
screen "704_Line_Overview_4" 1280x800
   Button "Button_19" at 852,670 size 37x32; TextOff 'Text'
      on Release: ActivateScreen("711_CARRIER_STATUS", 0)
      on Press: SetTag("HMI_EMS_Nr", "CarrierNumber")
   Button "Template_Button_3" at 1074,2 size 203x55; TextOn 'FAULT RESET FAULT RESET'; TextOff 'FAULT RESET FAULT RESET'
      on Release: ResetBit("DB_SDC_GLOBAL_M.SDC_ER_Reset")
      on Press: SetBit("DB_SDC_GLOBAL_M.SDC_ER_Reset")
   AlarmView "Template_Alarm view_2" at 128,2 size 948x112
   Button "Template_Button_4" at 1196,56 size 81x59; TextOff 'Text'
      Appearance <- "AlwaysTRUE"
   Button "Button_7" at 0,57 size 128x58; TextOff 'SELECT SCREEN'
      on Release: ActivateScreen("010_START", 0)
   Button "Button_6" at 0,0 size 128x58; TextOff 'PREVIOUS SCREEN'
      on Click: function_efd93a16()
   DateTimeField "Template_Date/time field_2" at 1075,56 size 123x28
   DateTimeField "Template_Date/time field_3" at 1075,83 size 122x32
   TextField "Text field_2" at 485,123 size 327x28; Text 'OVERVIEW 4 - SCREEN 704'
   GraphicView "Graphic view_1" at 439,169 size 432x627; Picture "Graphic_4"
   TextField "Text field_34" at 898,673 size 46x25; Text 'S34'
   TextField "Text field_93" at 584,373 size 60x24; Text 'EMS01'
   TextField "Text field_95" at 578,408 size 71x22; Text 'AREA E'
   Button "Button_2" at 988,687 size 127x87; TextOn 'LINE_OVERVIEW_2 LINE OVERVIEW_2'; TextOff 'LINE_OVERVIEW_2 System Overview Screen'
      on Click: ActivateScreen("700_System_Line_Overview", 0)
   Button "Button_1" at 1125,687 size 127x87; TextOn 'LINE_OVERVIEW_2 LINE OVERVIEW_2'; TextOff 'LINE_OVERVIEW_2 / Main Screen'
      on Click: ActivateScreen("010_START", 0)
   Button "Button_3" at 852,182 size 37x32; TextOff 'Text'
      on Release: ActivateScreen("711_CARRIER_STATUS", 0)
      on Press: SetTag("HMI_EMS_Nr", "CarrierNumber")
   Button "Button_4" at 852,215 size 37x32; TextOff 'Text'
      on Release: ActivateScreen("711_CARRIER_STATUS", 0)
      on Press: SetTag("HMI_EMS_Nr", "CarrierNumber")
   Button "Button_5" at 852,250 size 37x32; TextOff 'Text'
      on Release: ActivateScreen("711_CARRIER_STATUS", 0)
      on Press: SetTag("HMI_EMS_Nr", "CarrierNumber")
   Button "Button_8" at 852,285 size 37x32; TextOff 'Text'
      on Release: ActivateScreen("711_CARRIER_STATUS", 0)
      on Press: SetTag("HMI_EMS_Nr", "CarrierNumber")
   Button "Button_9" at 852,320 size 37x32; TextOff 'Text'
      on Release: ActivateScreen("711_CARRIER_STATUS", 0)
      on Press: SetTag("HMI_EMS_Nr", "CarrierNumber")
   Button "Button_10" at 852,355 size 37x32; TextOff 'Text'
      on Release: ActivateScreen("711_CARRIER_STATUS", 0)
      on Press: SetTag("HMI_EMS_Nr", "CarrierNumber")
   Button "Button_11" at 852,390 size 37x32; TextOff 'Text'
      on Release: ActivateScreen("711_CARRIER_STATUS", 0)
      on Press: SetTag("HMI_EMS_Nr", "CarrierNumber")
   Button "Button_12" at 852,425 size 37x32; TextOff 'Text'
      on Release: ActivateScreen("711_CARRIER_STATUS", 0)
      on Press: SetTag("HMI_EMS_Nr", "CarrierNumber")
   Button "Button_13" at 852,460 size 37x32; TextOff 'Text'
      on Release: ActivateScreen("711_CARRIER_STATUS", 0)
      on Press: SetTag("HMI_EMS_Nr", "CarrierNumber")
   Button "Button_14" at 852,495 size 37x32; TextOff 'Text'
      on Release: ActivateScreen("711_CARRIER_STATUS", 0)
      on Press: SetTag("HMI_EMS_Nr", "CarrierNumber")
   Button "Button_15" at 852,530 size 37x32; TextOff 'Text'
      on Release: ActivateScreen("711_CARRIER_STATUS", 0)
      on Press: SetTag("HMI_EMS_Nr", "CarrierNumber")
   Button "Button_16" at 852,565 size 37x32; TextOff 'Text'
      on Release: ActivateScreen("711_CARRIER_STATUS", 0)
      on Press: SetTag("HMI_EMS_Nr", "CarrierNumber")
   Button "Button_17" at 852,600 size 37x32; TextOff 'Text'
      on Release: ActivateScreen("711_CARRIER_STATUS", 0)
      on Press: SetTag("HMI_EMS_Nr", "CarrierNumber")
   Button "Button_18" at 852,635 size 37x32; TextOff 'Text'
      on Release: ActivateScreen("711_CARRIER_STATUS", 0)
      on Press: SetTag("HMI_EMS_Nr", "CarrierNumber")
   IOField "I/O field_50" at 852,670 size 37x32; FormatPattern 99
      ProcessValue <- "CarrierNumber"
      Appearance <- "Faulted"
   IOField "I/O field_32" at 852,182 size 37x32; FormatPattern 99
      ProcessValue <- "CarrierNumber"
      Appearance <- "Faulted"
   IOField "I/O field_33" at 852,215 size 37x32; FormatPattern 99
      ProcessValue <- "CarrierNumber"
      Appearance <- "Faulted"
   IOField "I/O field_34" at 852,250 size 37x32; FormatPattern 99
      ProcessValue <- "CarrierNumber"
      Appearance <- "Faulted"
   IOField "I/O field_35" at 852,285 size 37x32; FormatPattern 99
      ProcessValue <- "CarrierNumber"
      Appearance <- "Faulted"
   IOField "I/O field_36" at 852,320 size 37x32; FormatPattern 99
      ProcessValue <- "CarrierNumber"
      Appearance <- "Faulted"
   IOField "I/O field_49" at 852,635 size 37x32; FormatPattern 99
      ProcessValue <- "CarrierNumber"
      Appearance <- "Faulted"
   IOField "I/O field_40" at 852,600 size 37x32; FormatPattern 99
      ProcessValue <- "CarrierNumber"
      Appearance <- "Faulted"
   IOField "I/O field_41" at 852,565 size 37x32; FormatPattern 99
      ProcessValue <- "CarrierNumber"
      Appearance <- "Faulted"
   IOField "I/O field_43" at 852,530 size 37x32; FormatPattern 99
      ProcessValue <- "CarrierNumber"
      Appearance <- "Faulted"
   IOField "I/O field_44" at 852,495 size 37x32; FormatPattern 99
      ProcessValue <- "CarrierNumber"
      Appearance <- "Faulted"
   IOField "I/O field_45" at 852,460 size 37x32; FormatPattern 99
      ProcessValue <- "CarrierNumber"
      Appearance <- "Faulted"
   IOField "I/O field_46" at 852,425 size 37x32; FormatPattern 99
      ProcessValue <- "CarrierNumber"
      Appearance <- "Faulted"
   IOField "I/O field_47" at 852,390 size 37x32; FormatPattern 99
      ProcessValue <- "CarrierNumber"
      Appearance <- "Faulted"
   IOField "I/O field_48" at 852,355 size 37x32; FormatPattern 99
      ProcessValue <- "CarrierNumber"
      Appearance <- "Faulted"

screen "711_CARRIER_STATUS" 1280x800, template "Top_Header"
   on GenerateScreen: "SDC_EMS_STATUS"("HMI_EMS_Nr"); "SDC_EMS_TA_STATUS"("HMI_EMS_Nr"); "SDC_ERRORS"("HMI_EMS_Nr"); SetTag("SDC\DB_SDC_EMS\HMI[XX].BILD_Nr", 711); SetTag("SDC\_intern_Bildnummer", 711); "SDC_TS_REFERENCE"("SDC\DB_SDC_EMS\EMS[XXX].TS_STAT.VAL.SEK"); "SDC_GLOBAL_REFERENCE_PROFIL"("SDC\DB_SDC_EMS\EMS[XXX].PROFIL")
   on ClearScreen: SetTag("SDC\DB_SDC_EMS\HMI[XX].BILD_Nr", 0)
   IOField "EA-Feld_4" at 270,148 size 56x32; FormatPattern 99
      on OnFinishInput: "SDC_EMS_STATUS"("HMI_EMS_Nr"); "SDC_EMS_TA_STATUS"("HMI_EMS_Nr"); "SDC_ERRORS"("HMI_EMS_Nr")
      ProcessValue <- "HMI_EMS_Nr"
   TextField "Textfeld_3" at 378,151 size 118x25; Text 'EMS-No. / EMS-Number / Carrier-Number'
   Button "Schaltfläche_1" at 327,149 size 40x32; TextOff '+'
      on Click: function_dd21b452("HMI_EMS_Nr", 1); "SDC_EMS_STATUS"("HMI_EMS_Nr"); "SDC_EMS_TA_STATUS"("HMI_EMS_Nr"); "SDC_ERRORS"("HMI_EMS_Nr")
   Button "Schaltfläche_3" at 231,148 size 39x32; TextOff '-'
      on Click: function_b9b71300("HMI_EMS_Nr", 1); "SDC_EMS_STATUS"("HMI_EMS_Nr"); "SDC_EMS_TA_STATUS"("HMI_EMS_Nr"); "SDC_ERRORS"("HMI_EMS_Nr")
   IOField "EA-Feld_5" at 740,309 size 96x32; Authorization "Benutzerverwaltung"; FormatPattern 99999
      ProcessValue <- "HMI_Carrier_ActualSpeed"
   TextField "Textfeld_4" at 706,289 size 187x25; Text 'drive stop position [mm] / Drive Stopposition mm / Current Carrier Speed'
   Group "Gruppe" at 176,202 size 1068x49
   IOField "EA-Feld_14" at 788,216 size 48x28; FormatPattern 999
      on OnFinishInput: "SDC_EMS_STATUS"("HMI_EMS_Nr"); "SDC_TS_REFERENCE"("SDC\DB_SDC_EMS\EMS[XXX].TS_STAT.VAL.SEK"); "SDC_EMS_TA_STATUS"("HMI_EMS_Nr"); "SDC_ERRORS"("HMI_EMS_Nr")
      ProcessValue <- "HMI_EMS_Nr"
   IOField "EA-Feld_15" at 788,216 size 48x28; FormatPattern 999
      on OnFinishInput: "SDC_TS_PARAMETER"()
      Visibility <- "SDC\DB_SDC_EMS\EMS[XXX].TS_STAT.VAL.ERROR"
      ProcessValue <- "DB401_HMI_Status_CarrierFaultCode"
   TextField "Textfeld_17" at 726,216 size 50x22; Text 'ERROR / Error'
      Visibility <- "SDC\DB_SDC_EMS\EMS[XXX].ERRORS_SDC"
   IOField "EA-Feld_22" at 754,168 size 96x32; Authorization "Benutzerverwaltung"; FormatPattern 9999999999
      ProcessValue <- "HMI_Carrier_CurrentPosition"
   TextField "Textfeld_26" at 736,150 size 175x25; Text 'drive in position / Drive in Position / Current carrier position'
   TextField "Textfeld_29" at 1028,255 size 200x25; Text 'distance to next EMS / distance to preceding EMS / Next Stop Position'
   TextField "Textfeld_47" at 452,266 size 177x25; Text 'drives forward / EMS move forward / Carrier Moving Forward'
   Circle "Kreis_22" at 431,272 size 15x15
      Appearance <- "HMI_Carrier_RunningFwd"
   TextField "Textfeld_55" at 452,288 size 176x25; Text 'drives backward / EMS move reward / Carrier Moving Reverse'
   Circle "Kreis_30" at 431,294 size 15x15
      Appearance <- "HMI_Carrier_RunningRev"
   TextField "Textfeld_56" at 452,309 size 179x25; Text 'drive in position / EMS Drive in Position / Carrier Drive in Position'
   Circle "Kreis_31" at 431,315 size 15x15
      Appearance <- "HMI_Carrier_AtCommandPosition"
   Button "Schaltfläche_15" at 11,710 size 117x84; TextOff 'I / O EDIT CARRIER I/O'
      on Click: ActivateScreen("712_CARRIER_IO", 0)
   TextField "Textfeld_7" at 567,118 size 243x27; Text 'section counter / min Barcode mm / Carrier Status'
   Rectangle "Rectangle_1" at 11,443 size 55x42
      Appearance <- "HMI_Carrier_DriveCommFault"
   TextField "Textfeld_8" at 71,450 size 155x25; Text 'EMS Notbetrieb Tilt / EMS VAC CLEAN / G120 D Drive Status'
   Rectangle "Rectangle_2" at 11,494 size 55x42
      Appearance <- "HMI_Carrier_EncoderCommFault"
   TextField "Textfeld_9" at 74,501 size 148x25; Text 'EMS Notbetrieb Tilt / EMS VAC CLEAN / PnF Encoder Status'
   Rectangle "Rectangle_9" at 11,547 size 55x42
      Appearance <- "HMI_Carrier_HMICommFault"
   TextField "Textfeld_16" at 76,552 size 152x25; Text 'EMS Notbetrieb Tilt / EMS VAC CLEAN / IRD 400 HMI Status'
   TextField "Textfeld_19" at 12,400 size 242x26; Text 'EMS Notbetrieb Tilt / EMS VAC CLEAN / CARRIER DEVICE STATUS'
   Button "Schaltfläche_2" at 546,476 size 27x27; TextOff 'Text'; Authorization "Bedienen"
      on Click: function_c82f6f27("SDC\DB_SDC_EMS\EMS[XXX].FKT_SET", 8)
      ObjectEnable <- "SDC\DB_SDC_EMS\HMI[XX].FR_EDIT"
      Appearance <- "HMI_Carrier_Comm_Fault"
   Button "Schaltfläche_5" at 546,506 size 27x27; TextOff 'Text'; Authorization "Bedienen"
      on Click: function_c82f6f27("SDC\DB_SDC_EMS\EMS[XXX].FKT_SET", 10)
      ObjectEnable <- "SDC\DB_SDC_EMS\HMI[XX].FR_EDIT"
      Appearance <- "HMI_Carrier_Auto"
   Button "Schaltfläche_6" at 546,566 size 27x27; TextOff 'Text'; Authorization "Bedienen"
      on Click: function_c82f6f27("SDC\DB_SDC_EMS\EMS[XXX].FKT_SET", 12)
      ObjectEnable <- "SDC\DB_SDC_EMS\HMI[XX].FR_EDIT"
      Appearance <- "HMI_Carrier_Faulted"
   Button "Schaltfläche_7" at 546,596 size 27x27; TextOff 'Text'; Authorization "Bedienen"
      on Click: function_c82f6f27("SDC\DB_SDC_EMS\EMS[XXX].FKT_SET", 13)
      ObjectEnable <- "SDC\DB_SDC_EMS\HMI[XX].FR_EDIT"
      Appearance <- "HMI_Carrier_HoldPBPressed"
   Button "Schaltfläche_9" at 546,536 size 27x27; TextOff 'Text'; Authorization "Bedienen"
      on Click: function_c82f6f27("SDC\DB_SDC_EMS\EMS[XXX].FKT_SET", 11)
      ObjectEnable <- "SDC\DB_SDC_EMS\HMI[XX].FR_EDIT"
      Appearance <- "HMI_Carrier_Manual"
   TextField "Textfeld_59" at 579,598 size 176x25; Text 'Kohle Test n.i.O. / EMS TO REPAIR / CARRIER PROD. HOLD'
   TextField "Textfeld_1" at 579,507 size 148x25; Text 'EMS Notbetrieb Tilt / EMS VAC CLEAN / CARRIER IN AUTO'
   TextField "Textfeld_2" at 579,568 size 159x25; Text 'SMGM Qualität n.i.O. / EMS TO REPAIR / CARRIER FAULT'
   TextField "Textfeld_20" at 580,476 size 181x25; Text 'EMS Notbetrieb Tilt / EMS VAC CLEAN / CARRIER COMM FAULT'
   TextField "Textfeld_6" at 580,536 size 166x25; Text 'EMS Notbetrieb Tilt / EMS VAC CLEAN / CARRIER IN MANUAL'
   TextField "Textfeld_38" at 218,274 size 188x25; Text 'command drive forward / Command forward / Command Drive Forward'
   Circle "Kreis_13" at 194,280 size 15x15
      Appearance <- "HMI_Carrier_DriveFwdCommand"
   TextField "Textfeld_40" at 218,305 size 193x25; Text 'command drive backward / Command reward / Command Speed'
   IOField "EA-Feld_1" at 138,302 size 96x32; Authorization "Benutzerverwaltung"; FormatPattern 99999
      ProcessValue <- "HMI_Carrier_DriveCmdSpeed"
   Button "Schaltfläche_10" at 154,710 size 117x84; TextOff 'I / O EDIT CARRIER DRIVE'
      on Click: ActivateScreen("728_CARRIER_VFD_STATUS", 0)
   Button "Schaltfläche_11" at 300,710 size 117x84; TextOff 'I / O EDIT CARRIER FAULTS'
      on Click: ActivateScreen("713_CARRIER_FAULT", 0)
   IOField "EA-Feld_2" at 1116,273 size 96x32; Authorization "Benutzerverwaltung"; FormatPattern 99999999
      ProcessValue <- "HMI_Carrier_NextStopPosition"
   TextField "Textfeld_11" at 1030,147 size 200x25; Text 'distance to next EMS / distance to preceding EMS / Next Carrier Number'
   IOField "EA-Feld_3" at 1118,165 size 96x32; Authorization "Benutzerverwaltung"; FormatPattern 99999
      ProcessValue <- "HMI_Carrier_NextCarrierNumber"
   IOField "EA-Feld_30" at 951,487 size 56x32; FormatPattern 99
      on OnFinishInput: "SDC_TS_PARAMETER"()
      ProcessValue <- "HMI_Carrier_CurrentZone"
   TextField "Textfeld_37" at 825,487 size 174x27; Text 'section no. / Tracksectionnumber / Zone Number'
   TextField "Textfeld_5" at 825,466 size 174x27; Text 'section no. / Tracksectionnumber / Carrier in'
   Button "Schaltfläche_4" at 1089,543 size 117x84; TextOff 'I / O EDIT SET MASK CARRIER FAULTS'
      Appearance <- "Mask_Carrier_Faults_LT"
      on Press: SetBit("Set_Mask_Carrier_Faults_PB")
      on Release: ResetBit("Set_Mask_Carrier_Faults_PB")
   Button "Schaltfläche_8" at 1089,670 size 117x84; TextOff 'I / O EDIT RESET MASK CARRIER FAULTS'
      on Press: SetBit("Reset_Mask_Carrier_Faults_PB")
      on Release: ResetBit("Reset_Mask_Carrier_Faults_PB")
   IOField "EA-Feld_6" at 951,552 size 56x32; FormatPattern ??
      on OnFinishInput: "SDC_TS_PARAMETER"()
      ProcessValue <- "HMI_Carrier_CurrentArea"
   TextField "Textfeld_10" at 825,552 size 174x27; Text 'section no. / Tracksectionnumber / Area Number'
   TextField "Textfeld_12" at 825,531 size 174x27; Text 'section no. / Tracksectionnumber / Carrier in'

screen "713_CARRIER_FAULT" 1280x800, template "Top_Header"
   on GenerateScreen: "SDC_EMS_STATUS"('SDC\_EMS_Nr'); "SDC_TS_REFERENCE"("SDC\_TS_Nr"); SetTag("SDC\_intern_Bildnummer", 712); "SDC_EMS_TA_STATUS"("HMI_EMS_Nr"); SetTag("SDC\_intern_Bildnummer", 712)
   on ClearScreen: SetTag("SDC\DB_SDC_EMS\HMI[XX].BILD_Nr", 0)
   IOField "EA-Feld_4" at 510,185 size 56x32; FormatPattern 9999
      on OnFinishInput: "SDC_EMS_STATUS"("HMI_EMS_Nr"); "SDC_EMS_TA_STATUS"("HMI_EMS_Nr"); "SDC_ERRORS"("HMI_EMS_Nr")
      ProcessValue <- "HMI_EMS_Nr"
   TextField "Textfeld_3" at 618,188 size 118x25; Text 'EMS-No. / EMS-Number / Carrier-Number'
   Button "Schaltfläche_1" at 567,185 size 40x32; TextOff '+'
      on Click: function_dd21b452("HMI_EMS_Nr", 1); "SDC_EMS_STATUS"("HMI_EMS_Nr"); "SDC_EMS_TA_STATUS"("HMI_EMS_Nr"); "SDC_ERRORS"("HMI_EMS_Nr")
   Button "Schaltfläche_3" at 470,185 size 39x32; TextOff '-'
      on Click: function_b9b71300("HMI_EMS_Nr", 1); "SDC_EMS_STATUS"("HMI_EMS_Nr"); "SDC_EMS_TA_STATUS"("HMI_EMS_Nr"); "SDC_ERRORS"("HMI_EMS_Nr")
   TextField "Textfeld_7" at 550,118 size 243x27; Text 'section counter / min Barcode mm / Carrier Fault'
   Button "Button_1" at 84,303 size 50x246; TextOff 'Text'
   TextField "Textfeld_11" at 137,309 size 293x25; Text 'EMS-No. / EMS-Number / FAULT 01 - CARRIER GENERAL FAULT'
   TextField "Textfeld_10" at 137,335 size 238x25; Text 'EMS-No. / EMS-Number / FAULT 02 - MOTION ON FAULT'
   TextField "Textfeld_13" at 137,361 size 245x25; Text 'EMS-No. / EMS-Number / FAULT 03 - MOTION OFF FAULT'
   TextField "Textfeld_14" at 137,387 size 288x25; Text 'EMS-No. / EMS-Number / FAULT 04 - CARRIER SPACING FAULT'
   TextField "Textfeld_15" at 137,412 size 248x25; Text 'EMS-No. / EMS-Number / FAULT 05 - DRIVE COMM FAULT'
   TextField "Textfeld_16" at 137,438 size 272x25; Text 'EMS-No. / EMS-Number / FAULT 06 - DRIVE GENERAL FAULT'
   TextField "Textfeld_17" at 137,464 size 275x25; Text 'EMS-No. / EMS-Number / FAULT 07 - ENCODER COMM FAULT'
   TextField "Textfeld_18" at 137,490 size 265x25; Text 'EMS-No. / EMS-Number / FAULT 08 - CRASH DETECT FAULT'
   Circle "Kreis_13" at 102,312 size 15x15
      Appearance <- "DB401_HMI_Status_CarrierFaultCode"
   Circle "Kreis_1" at 102,338 size 15x15
      Appearance <- "DB401_HMI_Status_CarrierFaultCode"
   Circle "Kreis_2" at 102,364 size 15x15
      Appearance <- "DB401_HMI_Status_CarrierFaultCode"
   Circle "Kreis_3" at 102,390 size 15x15
      Appearance <- "DB401_HMI_Status_CarrierFaultCode"
   Circle "Kreis_4" at 102,416 size 15x15
      Appearance <- "DB401_HMI_Status_CarrierFaultCode"
   Circle "Kreis_5" at 102,442 size 15x15
      Appearance <- "DB401_HMI_Status_CarrierFaultCode"
   Circle "Kreis_6" at 102,468 size 15x15
      Appearance <- "DB401_HMI_Status_CarrierFaultCode"
   Circle "Kreis_7" at 102,494 size 15x15
      Appearance <- "DB401_HMI_Status_CarrierFaultCode"
   TextField "Textfeld_1" at 137,516 size 337x25; Text 'EMS-No. / EMS-Number / FAULT 15 - DRIVE ERROR INTERNAL COMM'
   Circle "Kreis_8" at 102,520 size 15x15
      Appearance <- "DB401_HMI_Status_CarrierFaultCode"
   Button "Button_2" at 516,303 size 50x246; TextOff 'Text'
   TextField "Textfeld_2" at 569,309 size 326x25; Text 'EMS-No. / EMS-Number / FAULT 20 - DRIVE MOTOR OVERCURRENT'
   TextField "Textfeld_4" at 569,335 size 273x25; Text 'EMS-No. / EMS-Number / FAULT 23 - DRIVE UNDERVOLTAGE'
   TextField "Textfeld_5" at 569,361 size 261x25; Text 'EMS-No. / EMS-Number / FAULT 24 - DRIVE OVERVOLTAGE'
   TextField "Textfeld_6" at 569,387 size 349x25; Text 'EMS-No. / EMS-Number / FAULT 25 - DRIVE PWR MODULE NOT READY'
   TextField "Textfeld_8" at 569,412 size 294x25; Text 'EMS-No. / EMS-Number / FAULT 32 - DRIVE MOTOR OVERTEMP'
   TextField "Textfeld_9" at 569,438 size 302x25; Text 'EMS-No. / EMS-Number / FAULT 40 - CARRIER NUMBER INVALID'
   TextField "Textfeld_12" at 569,464 size 302x25; Text 'EMS-No. / EMS-Number / FAULT 60 - ENCODER POSITION FAULT'
   Circle "Kreis_9" at 534,312 size 15x15
      Appearance <- "DB401_HMI_Status_CarrierFaultCode"
   Circle "Kreis_10" at 534,338 size 15x15
      Appearance <- "DB401_HMI_Status_CarrierFaultCode"
   Circle "Kreis_11" at 534,364 size 15x15
      Appearance <- "DB401_HMI_Status_CarrierFaultCode"
   Circle "Kreis_12" at 534,390 size 15x15
      Appearance <- "DB401_HMI_Status_CarrierFaultCode"
   Circle "Kreis_14" at 534,416 size 15x15
      Appearance <- "DB401_HMI_Status_CarrierFaultCode"
   Circle "Kreis_15" at 534,442 size 15x15
      Appearance <- "DB401_HMI_Status_CarrierFaultCode"
   Circle "Kreis_16" at 534,468 size 15x15
      Appearance <- "DB401_HMI_Status_CarrierFaultCode"
   TextField "Textfeld_20" at 569,489 size 339x25; Text 'EMS-No. / EMS-Number / FAULT DUP - DUPLICATE CARRIER # FAULT'
   Circle "Kreis_18" at 534,493 size 15x15
      Appearance <- "DB401_HMI_Status_CarrierFaultCode"

screen "715_ACCESS_POINT_LAYOUT" 1280x800
   GraphicView "Graphic view_1" at 0,119 size 1144x681; Picture "LAYOUT 1"
   Button "Button_9" at 451,171 size 47x26; TextOff 'AP6'
      Appearance <- "[106]"
   Button "Button_12" at 517,123 size 46x26; TextOff 'AP7'
      Appearance <- "[107]"
   Button "Button_10" at 574,123 size 46x26; TextOff 'AP8'
      Appearance <- "[108]"
   Button "Button_11" at 627,123 size 45x26; TextOff 'AP9'
      Appearance <- "[109]"
   Button "Button_13" at 694,171 size 47x26; TextOff 'AP5'
      Appearance <- "[105]"
   Button "Button_8" at 734,123 size 50x26; TextOff 'AP10'
      Appearance <- "[110]"
   Button "Button_14" at 749,222 size 52x26; TextOff 'AP11'
      Appearance <- "[111]"
   Button "Button_7" at 750,325 size 51x26; TextOff 'AP4'
      Appearance <- "[104]"
   Button "Button_6" at 749,444 size 52x26; TextOff 'AP12'
      Appearance <- "[112]"
   Button "Button_5" at 751,607 size 51x26; TextOff 'AP3'
      Appearance <- "[103]"
   Button "Button_4" at 777,637 size 52x26; TextOff 'AP13'
      Appearance <- "[113]"
   Button "Button_15" at 576,726 size 52x26; TextOff 'AP14'
      Appearance <- "[114]"
   Button "Button_16" at 384,711 size 53x26; TextOff 'AP15'
      Appearance <- "[115]"
   Button "Button_17" at 295,743 size 52x26; TextOff 'AP16'
      Appearance <- "[116]"
   Button "Button_18" at 267,687 size 53x26; TextOff 'AP17'
      Appearance <- "[117]"
   Button "Button_19" at 329,611 size 51x26; TextOff 'AP18'
      Appearance <- "[118]"
   Button "Button_1" at 479,611 size 50x26; TextOff 'AP1'
      Appearance <- "[101]"
   Button "Button_2" at 620,612 size 50x26; TextOff 'AP2'
      Appearance <- "[102]"
   TextField "Text field_126" at 847,138 size 369x28; Text 'ACCESS POINT LAYOUT SCREEN'
   Button "Button_20" at 471,117 size 46x26; TextOff 'AP19'
      Appearance <- "[119]"
   Button "Template_Button_3" at 1074,2 size 203x55; TextOn 'FAULT RESET FAULT RESET'; TextOff 'FAULT RESET FAULT RESET'
      on Release: ResetBit("DB_SDC_GLOBAL_M.SDC_ER_Reset")
      on Press: SetBit("DB_SDC_GLOBAL_M.SDC_ER_Reset")
   AlarmView "Template_Alarm view_2" at 128,2 size 948x112
   Button "Template_Button_4" at 1196,56 size 81x59; TextOff 'Text'
      Appearance <- "AlwaysTRUE"
   Button "Button_21" at 0,57 size 128x58; TextOff 'SELECT SCREEN'
      on Release: ActivateScreen("010_START", 0)
   Button "Button_22" at 0,0 size 128x58; TextOff 'PREVIOUS SCREEN'
      on Click: function_efd93a16()
   DateTimeField "Template_Date/time field_2" at 1075,56 size 123x28
   DateTimeField "Template_Date/time field_3" at 1075,83 size 122x32

screen "708_ZONE_STATUS" 1280x800, template "Top_Header"
   on GenerateScreen: "SDC_TS_PARAMETER"(); "SDC_TS_REFERENCE"("HMI_Zone_Nr"); SetTag("SDC\DB_SDC_TS_PARAMETER\DB_SDC_TS_PARAMETER_HMI.HMI[XX].BILD_Nr", 704); SetTag("SDC\_intern_Bildnummer", 704)
   on ClearScreen: SetTag("SDC\DB_SDC_TS_PARAMETER\DB_SDC_TS_PARAMETER_HMI.HMI[XX].BILD_Nr", 0)
   IOField "EA-Feld_1" at 144,392 size 96x32; Authorization "Benutzerverwaltung"; FormatPattern 9999999999
      Appearance <- "SDC\DB_SDC_TS_PARAMETER\DB_SDC_TS_PARAMETER_HMI.HMI[XX].FR_EDIT"
      ObjectEnable <- "SDC\DB_SDC_TS_PARAMETER\DB_SDC_TS_PARAMETER_HMI.HMI[XX].FR_EDIT"
      ProcessValue <- "DB401_HMI_Status_ZoneStatus.ZoneStartPosition"
   TextField "Textfeld_1" at 137,344 size 272x58; Text 'barcode value at start of section [mm] Sektion Start Barcode mm Position at start of zone [mm]'
   IOField "EA-Feld_2" at 1022,324 size 96x32; Authorization "Benutzerverwaltung"; FormatPattern 9999999999
      Appearance <- "SDC\DB_SDC_TS_PARAMETER\DB_SDC_TS_PARAMETER_HMI.HMI[XX].FR_EDIT"
      ObjectEnable <- "SDC\DB_SDC_TS_PARAMETER\DB_SDC_TS_PARAMETER_HMI.HMI[XX].FR_EDIT"
      ProcessValue <- "DB401_HMI_Status_ZoneStatus.ZoneEndPosition"
   TextField "Textfeld_2" at 743,318 size 275x59; Text 'barcode value at end of section [mm] Sektion Ende Barcode mm Position at end of zone [mm]'
   IOField "EA-Feld_4" at 416,188 size 56x32; FormatPattern 9999
      on OnFinishInput: "SDC_TS_PARAMETER"(); "SDC_TS_REFERENCE"("HMI_Zone_Nr")
      ProcessValue <- "HMI_Zone_Nr"
   TextField "Textfeld_3" at 515,188 size 93x33; Text 'section no. / Sektionnumber / Zone No'
   Button "Schaltfläche_1" at 473,188 size 40x32; TextOff '+'
      on Click: function_dd21b452("HMI_Zone_Nr", 1); "SDC_TS_PARAMETER"(); "SDC_TS_REFERENCE"("HMI_Zone_Nr")
   Button "Schaltfläche_3" at 376,188 size 39x32; TextOff '-'
      on Click: function_b9b71300("HMI_Zone_Nr", 1); "SDC_TS_PARAMETER"(); "SDC_TS_REFERENCE"("HMI_Zone_Nr")
   IOField "EA-Feld_8" at 1056,188 size 56x32; Authorization "Benutzerverwaltung"; FormatPattern 9999
      Appearance <- "SDC\DB_SDC_TS_PARAMETER\DB_SDC_TS_PARAMETER_HMI.HMI[XX].FR_EDIT"
      ObjectEnable <- "SDC\DB_SDC_TS_PARAMETER\DB_SDC_TS_PARAMETER_HMI.HMI[XX].FR_EDIT"
      ProcessValue <- "DB401_HMI_Status_ZoneStatus.NextZoneNumber"
   TextField "Textfeld_7" at 957,187 size 107x33; Text 'next section 1 / next Sektion 1 / Next Zone'
   Group "Gruppe" at 141,244 size 1024x49
   IOField "EA-Feld_13" at 610,192 size 163x24; Authorization "Benutzerverwaltung"; FormatPattern ????????????????
      Appearance <- "SDC\DB_SDC_TS_PARAMETER\DB_SDC_TS_PARAMETER_HMI.HMI[XX].FR_EDIT"
      ObjectEnable <- "SDC\DB_SDC_TS_PARAMETER\DB_SDC_TS_PARAMETER_HMI.HMI[XX].FR_EDIT"
      ProcessValue <- "DB401_HMI_Status_ZoneStatus.ZoneType"
   TextField "Textfeld_5" at 658,381 size 330x33; Text 'stop position (offset start) mm / Stopposition (Offset Start) mm / Zone Full'
   TextField "Textfeld_6" at 659,422 size 330x33; Text 'stop position (offset start) mm / Stopposition (Offset Start) mm / Speed Zone'
   TextField "Textfeld_8" at 659,463 size 330x33; Text 'stop position (offset start) mm / Stopposition (Offset Start) mm / Speed Zone Start'
   TextField "Textfeld_9" at 659,504 size 330x33; Text 'stop position (offset start) mm / Stopposition (Offset Start) mm / Speed Zone End'
   IOField "EA-Feld_3" at 596,460 size 56x32; FormatPattern 9999999999
      on OnFinishInput: "SDC_TS_PARAMETER"(); "SDC_TS_REFERENCE"("SDC\_TS_Nr")
      ProcessValue <- "DB401_HMI_Status_ZoneStatus.SpeedZoneStartPos"
   IOField "EA-Feld_6" at 596,500 size 56x32; FormatPattern 9999999999
      on OnFinishInput: "SDC_TS_PARAMETER"(); "SDC_TS_REFERENCE"("SDC\_TS_Nr")
      ProcessValue <- "DB401_HMI_Status_ZoneStatus.SpeedZoneEndPos"
   Circle "Kreis_13" at 616,387 size 15x15
      Appearance <- "DB401_HMI_Status_ZoneStatus.ZoneFull"
   Circle "Kreis_1" at 616,427 size 15x15
      Appearance <- "DB401_HMI_Status_ZoneStatus.SpeedZone"
   IOField "EA-Feld_9" at 596,540 size 56x32; Authorization "Benutzerverwaltung"; FormatPattern 99999
      Appearance <- "SDC\DB_SDC_TS_PARAMETER\DB_SDC_TS_PARAMETER_HMI.HMI[XX].FR_EDIT"
      ObjectEnable <- "SDC\DB_SDC_TS_PARAMETER\DB_SDC_TS_PARAMETER_HMI.HMI[XX].FR_EDIT"
      ProcessValue <- "DB401_HMI_Status_ZoneStatus.AccumZoneSpacing"
   TextField "Textfeld_11" at 659,542 size 330x33; Text 'stop position (offset start) mm / Stopposition (Offset Start) mm / Accum Zone Spacing'
   IOField "EA-Feld_10" at 596,580 size 56x32; Authorization "Benutzerverwaltung"; FormatPattern 99999
      Appearance <- "SDC\DB_SDC_TS_PARAMETER\DB_SDC_TS_PARAMETER_HMI.HMI[XX].FR_EDIT"
      ObjectEnable <- "SDC\DB_SDC_TS_PARAMETER\DB_SDC_TS_PARAMETER_HMI.HMI[XX].FR_EDIT"
      ProcessValue <- "DB401_HMI_Status_ZoneStatus.ProductionZoneSpacing"
   TextField "Textfeld_12" at 659,582 size 330x33; Text 'stop position (offset start) mm / Stopposition (Offset Start) mm / Prooduction Zone Spacing'
   TextField "Textfeld_13" at 459,114 size 243x27; Text 'section counter / min Barcode mm / Zone Status'
   TextField "Text field_1" at 911,358 size 101x25; Text 'Stop Position'
   TextField "Text field_2" at 642,168 size 83x25; Text 'Zone Type'
   IOField "EA-Feld_5" at 119,189 size 56x32; Authorization "Benutzerverwaltung"; FormatPattern 9999
      Appearance <- "SDC\DB_SDC_TS_PARAMETER\DB_SDC_TS_PARAMETER_HMI.HMI[XX].FR_EDIT"
      ObjectEnable <- "SDC\DB_SDC_TS_PARAMETER\DB_SDC_TS_PARAMETER_HMI.HMI[XX].FR_EDIT"
      ProcessValue <- "DB401_HMI_Status_ZoneStatus.PrevZoneNumber"
   TextField "Textfeld_4" at 25,189 size 94x33; Text 'next section 1 / next Sektion 1 / Prev Zone'

VB script "SDC_EMS_FLAGS"
   'HINWEIS:
   ' Beim Erstellen von Skripten können Sie mit <Strg+Leertaste> vordefinierte 
   ' Systemfunktionen in das neue Skript einbinden.
   ' Das HMIRuntime-Objekt ermöglicht einfachen Zugriff auf die Objekte des
   ' WinCC flexible Objektmodells, ihre Methoden und ihre Eigenschaften.
   ' Für ein komfortables Auswählen einer Objektreferenz betätigen Sie bitte <Alt+Rechts>.
   ' Komplexe Skripte können Sie mit Sprachelementen der Programmiersprache
   ' VBScript erstellen.
   ' Der Zugriff auf WinCC flexible Variablen erfolgt direkt über den Variablennamen,
   ' z.B. Tag = 5
   
   '________________________________________________________________________________
   '
   
   ' Groiß Andreas
   ' Siemens AG Österreich 
   ' Linz Kraußstraße 1-7 
   ' RC-AT I-IA AS-FA-SO-AE2
   ' 28.01.2015
   
   Dim EMS_Nr ' Sektion Number
   Dim Laenge_Data ' Länge FLAG Daten
   Dim Allg_Offset ' Allg Parameter Offset
   Dim HMIFlagDaten_Offset ' HMI Sektionsdaten Offset
   Dim HMI_Nr ' HMI Nummer
   
   ' INIT-------------------------------------------------------------
   
   If (SmartTags("SDC\DB_SDC_EMS_FLAGS\_EMS_Nr") < SmartTags("DB_SDC_GLOBAL_EMS_ID_MIN")) Or (SmartTags("SDC\DB_SDC_EMS_FLAGS\_EMS_Nr") > SmartTags("DB_SDC_GLOBAL_EMS_ID_MAX")) Then
   	SmartTags("SDC\DB_SDC_EMS_FLAGS\_EMS_Nr") = 	SmartTags("DB_SDC_GLOBAL_EMS_ID_MIN")
   End If	
   
   If (SmartTags("SDC\DB_SDC_EMS_FLAGS\_EMS_Nr") < 1) Then
   	SmartTags("SDC\DB_SDC_EMS_FLAGS\_EMS_Nr") = 1
   End If	
   
   '##############################################
   ' S7 sucht sich Daten:
   '##############################################
   
       Laenge_Data = SmartTags("DB_SDC_EMS_FLAGS_HEADER.LAENGE_EMS_FLAGS")
       Allg_Offset = SmartTags("DB_SDC_EMS_FLAGS_HEADER.START_EMS")
   
       SmartTags("SDC\DB_SDC_EMS_FLAGS\_EMS_Flags_Byte_EMS001") = 001 * Laenge_Data - Laenge_Data + Allg_Offset 
       SmartTags("SDC\DB_SDC_EMS_FLAGS\_EMS_Flags_Byte_EMS002") = 002 * Laenge_Data - Laenge_Data + Allg_Offset 
       SmartTags("SDC\DB_SDC_EMS_FLAGS\_EMS_Flags_Byte_EMS003") = 003 * Laenge_Data - Laenge_Data + Allg_Offset 
       SmartTags("SDC\DB_SDC_EMS_FLAGS\_EMS_Flags_Byte_EMS004") = 004 * Laenge_Data - Laenge_Data + Allg_Offset 
       SmartTags("SDC\DB_SDC_EMS_FLAGS\_EMS_Flags_Byte_EMS005") = 005 * Laenge_Data - Laenge_Data + Allg_Offset 
       SmartTags("SDC\DB_SDC_EMS_FLAGS\_EMS_Flags_Byte_EMS006") = 006 * Laenge_Data - Laenge_Data + Allg_Offset 
       SmartTags("SDC\DB_SDC_EMS_FLAGS\_EMS_Flags_Byte_EMS007") = 007 * Laenge_Data - Laenge_Data + Allg_Offset 
       SmartTags("SDC\DB_SDC_EMS_FLAGS\_EMS_Flags_Byte_EMS008") = 008 * Laenge_Data - Laenge_Data + Allg_Offset 
       SmartTags("SDC\DB_SDC_EMS_FLAGS\_EMS_Flags_Byte_EMS009") = 009 * Laenge_Data - Laenge_Data + Allg_Offset 
       SmartTags("SDC\DB_SDC_EMS_FLAGS\_EMS_Flags_Byte_EMS010") = 010 * Laenge_Data - Laenge_Data + Allg_Offset 
       SmartTags("SDC\DB_SDC_EMS_FLAGS\_EMS_Flags_Byte_EMS011") = 011 * Laenge_Data - Laenge_Data + Allg_Offset 
       SmartTags("SDC\DB_SDC_EMS_FLAGS\_EMS_Flags_Byte_EMS012") = 012 * Laenge_Data - Laenge_Data + Allg_Offset 
       SmartTags("SDC\DB_SDC_EMS_FLAGS\_EMS_Flags_Byte_EMS013") = 013 * Laenge_Data - Laenge_Data + Allg_Offset 
       SmartTags("SDC\DB_SDC_EMS_FLAGS\_EMS_Flags_Byte_EMS014") = 014 * Laenge_Data - Laenge_Data + Allg_Offset 
       SmartTags("SDC\DB_SDC_EMS_FLAGS\_EMS_Flags_Byte_EMS015") = 015 * Laenge_Data - Laenge_Data + Allg_Offset 
       SmartTags("SDC\DB_SDC_EMS_FLAGS\_EMS_Flags_Byte_EMS016") = 016 * Laenge_Data - Laenge_Data + Allg_Offset 
       SmartTags("SDC\DB_SDC_EMS_FLAGS\_EMS_Flags_Byte_EMS017") = 017 * Laenge_Data - Laenge_Data + Allg_Offset 
       SmartTags("SDC\DB_SDC_EMS_FLAGS\_EMS_Flags_Byte_EMS018") = 018 * Laenge_Data - Laenge_Data + Allg_Offset 
       SmartTags("SDC\DB_SDC_EMS_FLAGS\_EMS_Flags_Byte_EMS019") = 019 * Laenge_Data - Laenge_Data + Allg_Offset 
       SmartTags("SDC\DB_SDC_EMS_FLAGS\_EMS_Flags_Byte_EMS020") = 020 * Laenge_Data - Laenge_Data + Allg_Offset 
       SmartTags("SDC\DB_SDC_EMS_FLAGS\_EMS_Flags_Byte_EMS021") = 021 * Laenge_Data - Laenge_Data + Allg_Offset 
       SmartTags("SDC\DB_SDC_EMS_FLAGS\_EMS_Flags_Byte_EMS022") = 022 * Laenge_Data - Laenge_Data + Allg_Offset 
       SmartTags("SDC\DB_SDC_EMS_FLAGS\_EMS_Flags_Byte_EMS023") = 023 * Laenge_Data - Laenge_Data + Allg_Offset 
       SmartTags("SDC\DB_SDC_EMS_FLAGS\_EMS_Flags_Byte_EMS024") = 024 * Laenge_Data - Laenge_Data + Allg_Offset 
       SmartTags("SDC\DB_SDC_EMS_FLAGS\_EMS_Flags_Byte_EMS025") = 025 * Laenge_Data - Laenge_Data + Allg_Offset 
       SmartTags("SDC\DB_SDC_EMS_FLAGS\_EMS_Flags_Byte_EMS026") = 026 * Laenge_Data - Laenge_Data + Allg_Offset 
       SmartTags("SDC\DB_SDC_EMS_FLAGS\_EMS_Flags_Byte_EMS027") = 027 * Laenge_Data - Laenge_Data + Allg_Offset 
       SmartTags("SDC\DB_SDC_EMS_FLAGS\_EMS_Flags_Byte_EMS028") = 028 * Laenge_Data - Laenge_Data + Allg_Offset 
       SmartTags("SDC\DB_SDC_EMS_FLAGS\_EMS_Flags_Byte_EMS029") = 029 * Laenge_Data - Laenge_Data + Allg_Offset 
       SmartTags("SDC\DB_SDC_EMS_FLAGS\_EMS_Flags_Byte_EMS030") = 030 * Laenge_Data - Laenge_Data + Allg_Offset 
       SmartTags("SDC\DB_SDC_EMS_FLAGS\_EMS_Flags_Byte_EMS031") = 031 * Laenge_Data - Laenge_Data + Allg_Offset 
       SmartTags("SDC\DB_SDC_EMS_FLAGS\_EMS_Flags_Byte_EMS032") = 032 * Laenge_Data - Laenge_Data + Allg_Offset 
       SmartTags("SDC\DB_SDC_EMS_FLAGS\_EMS_Flags_Byte_EMS033") = 033 * Laenge_Data - Laenge_Data + Allg_Offset 
       SmartTags("SDC\DB_SDC_EMS_FLAGS\_EMS_Flags_Byte_EMS034") = 034 * Laenge_Data - Laenge_Data + Allg_Offset 
       SmartTags("SDC\DB_SDC_EMS_FLAGS\_EMS_Flags_Byte_EMS035") = 035 * Laenge_Data - Laenge_Data + Allg_Offset 
       SmartTags("SDC\DB_SDC_EMS_FLAGS\_EMS_Flags_Byte_EMS036") = 036 * Laenge_Data - Laenge_Data + Allg_Offset 
       SmartTags("SDC\DB_SDC_EMS_FLAGS\_EMS_Flags_Byte_EMS037") = 037 * Laenge_Data - Laenge_Data + Allg_Offset 
       SmartTags("SDC\DB_SDC_EMS_FLAGS\_EMS_Flags_Byte_EMS038") = 038 * Laenge_Data - Laenge_Data + Allg_Offset 
       SmartTags("SDC\DB_SDC_EMS_FLAGS\_EMS_Flags_Byte_EMS039") = 039 * Laenge_Data - Laenge_Data + Allg_Offset     
       SmartTags("SDC\DB_SDC_EMS_FLAGS\_EMS_Flags_Byte_EMS040") = 040 * Laenge_Data - Laenge_Data + Allg_Offset 
       SmartTags("SDC\DB_SDC_EMS_FLAGS\_EMS_Flags_Byte_EMS041") = 041 * Laenge_Data - Laenge_Data + Allg_Offset 
       SmartTags("SDC\DB_SDC_EMS_FLAGS\_EMS_Flags_Byte_EMS042") = 042 * Laenge_Data - Laenge_Data + Allg_Offset 
       SmartTags("SDC\DB_SDC_EMS_FLAGS\_EMS_Flags_Byte_EMS043") = 043 * Laenge_Data - Laenge_Data + Allg_Offset 
       SmartTags("SDC\DB_SDC_EMS_FLAGS\_EMS_Flags_Byte_EMS044") = 044 * Laenge_Data - Laenge_Data + Allg_Offset 
       SmartTags("SDC\DB_SDC_EMS_FLAGS\_EMS_Flags_Byte_EMS045") = 045 * Laenge_Data - Laenge_Data + Allg_Offset 
       SmartTags("SDC\DB_SDC_EMS_FLAGS\_EMS_Flags_Byte_EMS046") = 046 * Laenge_Data - Laenge_Data + Allg_Offset 
       SmartTags("SDC\DB_SDC_EMS_FLAGS\_EMS_Flags_Byte_EMS047") = 047 * Laenge_Data - Laenge_Data + Allg_Offset 
       SmartTags("SDC\DB_SDC_EMS_FLAGS\_EMS_Flags_Byte_EMS048") = 048 * Laenge_Data - Laenge_Data + Allg_Offset 
       SmartTags("SDC\DB_SDC_EMS_FLAGS\_EMS_Flags_Byte_EMS049") = 049 * Laenge_Data - Laenge_Data + Allg_Offset     
       SmartTags("SDC\DB_SDC_EMS_FLAGS\_EMS_Flags_Byte_EMS050") = 050 * Laenge_Data - Laenge_Data + Allg_Offset 
       SmartTags("SDC\DB_SDC_EMS_FLAGS\_EMS_Flags_Byte_EMS051") = 051 * Laenge_Data - Laenge_Data + Allg_Offset 
       SmartTags("SDC\DB_SDC_EMS_FLAGS\_EMS_Flags_Byte_EMS052") = 052 * Laenge_Data - Laenge_Data + Allg_Offset 
       SmartTags("SDC\DB_SDC_EMS_FLAGS\_EMS_Flags_Byte_EMS053") = 053 * Laenge_Data - Laenge_Data + Allg_Offset 
       SmartTags("SDC\DB_SDC_EMS_FLAGS\_EMS_Flags_Byte_EMS054") = 054 * Laenge_Data - Laenge_Data + Allg_Offset 
       SmartTags("SDC\DB_SDC_EMS_FLAGS\_EMS_Flags_Byte_EMS055") = 055 * Laenge_Data - Laenge_Data + Allg_Offset 
       SmartTags("SDC\DB_SDC_EMS_FLAGS\_EMS_Flags_Byte_EMS056") = 056 * Laenge_Data - Laenge_Data + Allg_Offset 
       SmartTags("SDC\DB_SDC_EMS_FLAGS\_EMS_Flags_Byte_EMS057") = 057 * Laenge_Data - Laenge_Data + Allg_Offset 
       SmartTags("SDC\DB_SDC_EMS_FLAGS\_EMS_Flags_Byte_EMS058") = 058 * Laenge_Data - Laenge_Data + Allg_Offset 
       SmartTags("SDC\DB_SDC_EMS_FLAGS\_EMS_Flags_Byte_EMS059") = 059 * Laenge_Data - Laenge_Data + Allg_Offset 
       SmartTags("SDC\DB_SDC_EMS_FLAGS\_EMS_Flags_Byte_EMS060") = 060 * Laenge_Data - Laenge_Data + Allg_Offset 
       SmartTags("SDC\DB_SDC_EMS_FLAGS\_EMS_Flags_Byte_EMS061") = 061 * Laenge_Data - Laenge_Data + Allg_Offset 
       SmartTags("SDC\DB_SDC_EMS_FLAGS\_EMS_Flags_Byte_EMS062") = 062 * Laenge_Data - Laenge_Data + Allg_Offset 
       SmartTags("SDC\DB_SDC_EMS_FLAGS\_EMS_Flags_Byte_EMS063") = 063 * Laenge_Data - Laenge_Data + Allg_Offset 
       SmartTags("SDC\DB_SDC_EMS_FLAGS\_EMS_Flags_Byte_EMS064") = 064 * Laenge_Data - Laenge_Data + Allg_Offset 
       SmartTags("SDC\DB_SDC_EMS_FLAGS\_EMS_Flags_Byte_EMS065") = 065 * Laenge_Data - Laenge_Data + Allg_Offset 
       SmartTags("SDC\DB_SDC_EMS_FLAGS\_EMS_Flags_Byte_EMS066") = 066 * Laenge_Data - Laenge_Data + Allg_Offset 
       SmartTags("SDC\DB_SDC_EMS_FLAGS\_EMS_Flags_Byte_EMS067") = 067 * Laenge_Data - Laenge_Data + Allg_Offset 
       SmartTags("SDC\DB_SDC_EMS_FLAGS\_EMS_Flags_Byte_EMS068") = 068 * Laenge_Data - Laenge_Data + Allg_Offset 
       SmartTags("SDC\DB_SDC_EMS_FLAGS\_EMS_Flags_Byte_EMS069") = 069 * Laenge_Data - Laenge_Data + Allg_Offset 
       SmartTags("SDC\DB_SDC_EMS_FLAGS\_EMS_Flags_Byte_EMS070") = 070 * Laenge_Data - Laenge_Data + Allg_Offset 
       SmartTags("SDC\DB_SDC_EMS_FLAGS\_EMS_Flags_Byte_EMS071") = 071 * Laenge_Data - Laenge_Data + Allg_Offset 
       SmartTags("SDC\DB_SDC_EMS_FLAGS\_EMS_Flags_Byte_EMS072") = 072 * Laenge_Data - Laenge_Data + Allg_Offset 
       SmartTags("SDC\DB_SDC_EMS_FLAGS\_EMS_Flags_Byte_EMS073") = 073 * Laenge_Data - Laenge_Data + Allg_Offset 
       SmartTags("SDC\DB_SDC_EMS_FLAGS\_EMS_Flags_Byte_EMS074") = 074 * Laenge_Data - Laenge_Data + Allg_Offset 
       SmartTags("SDC\DB_SDC_EMS_FLAGS\_EMS_Flags_Byte_EMS075") = 075 * Laenge_Data - Laenge_Data + Allg_Offset 
       SmartTags("SDC\DB_SDC_EMS_FLAGS\_EMS_Flags_Byte_EMS076") = 076 * Laenge_Data - Laenge_Data + Allg_Offset 
       SmartTags("SDC\DB_SDC_EMS_FLAGS\_EMS_Flags_Byte_EMS077") = 077 * Laenge_Data - Laenge_Data + Allg_Offset 
       SmartTags("SDC\DB_SDC_EMS_FLAGS\_EMS_Flags_Byte_EMS078") = 078 * Laenge_Data - Laenge_Data + Allg_Offset 
       SmartTags("SDC\DB_SDC_EMS_FLAGS\_EMS_Flags_Byte_EMS079") = 079 * Laenge_Data - Laenge_Data + Allg_Offset 
       SmartTags("SDC\DB_SDC_EMS_FLAGS\_EMS_Flags_Byte_EMS080") = 080 * Laenge_Data - Laenge_Data + Allg_Offset 
       SmartTags("SDC\DB_SDC_EMS_FLAGS\_EMS_Flags_Byte_EMS081") = 081 * Laenge_Data - Laenge_Data + Allg_Offset 
       SmartTags("SDC\DB_SDC_EMS_FLAGS\_EMS_Flags_Byte_EMS082") = 082 * Laenge_Data - Laenge_Data + Allg_Offset 
       SmartTags("SDC\DB_SDC_EMS_FLAGS\_EMS_Flags_Byte_EMS083") = 083 * Laenge_Data - Laenge_Data + Allg_Offset 
       SmartTags("SDC\DB_SDC_EMS_FLAGS\_EMS_Flags_Byte_EMS084") = 084 * Laenge_Data - Laenge_Data + Allg_Offset 
       SmartTags("SDC\DB_SDC_EMS_FLAGS\_EMS_Flags_Byte_EMS085") = 085 * Laenge_Data - Laenge_Data + Allg_Offset 
       SmartTags("SDC\DB_SDC_EMS_FLAGS\_EMS_Flags_Byte_EMS086") = 086 * Laenge_Data - Laenge_Data + Allg_Offset 
       SmartTags("SDC\DB_SDC_EMS_FLAGS\_EMS_Flags_Byte_EMS087") = 087 * Laenge_Data - Laenge_Data + Allg_Offset 
       SmartTags("SDC\DB_SDC_EMS_FLAGS\_EMS_Flags_Byte_EMS088") = 088 * Laenge_Data - Laenge_Data + Allg_Offset 
       SmartTags("SDC\DB_SDC_EMS_FLAGS\_EMS_Flags_Byte_EMS089") = 089 * Laenge_Data - Laenge_Data + Allg_Offset     
       SmartTags("SDC\DB_SDC_EMS_FLAGS\_EMS_Flags_Byte_EMS090") = 090 * Laenge_Data - Laenge_Data + Allg_Offset 
       SmartTags("SDC\DB_SDC_EMS_FLAGS\_EMS_Flags_Byte_EMS091") = 091 * Laenge_Data - Laenge_Data + Allg_Offset 
       SmartTags("SDC\DB_SDC_EMS_FLAGS\_EMS_Flags_Byte_EMS092") = 092 * Laenge_Data - Laenge_Data + Allg_Offset 
       SmartTags("SDC\DB_SDC_EMS_FLAGS\_EMS_Flags_Byte_EMS093") = 093 * Laenge_Data - Laenge_Data + Allg_Offset 
       SmartTags("SDC\DB_SDC_EMS_FLAGS\_EMS_Flags_Byte_EMS094") = 094 * Laenge_Data - Laenge_Data + Allg_Offset 
       SmartTags("SDC\DB_SDC_EMS_FLAGS\_EMS_Flags_Byte_EMS095") = 095 * Laenge_Data - Laenge_Data + Allg_Offset 
       SmartTags("SDC\DB_SDC_EMS_FLAGS\_EMS_Flags_Byte_EMS096") = 096 * Laenge_Data - Laenge_Data + Allg_Offset 
       SmartTags("SDC\DB_SDC_EMS_FLAGS\_EMS_Flags_Byte_EMS097") = 097 * Laenge_Data - Laenge_Data + Allg_Offset 
       SmartTags("SDC\DB_SDC_EMS_FLAGS\_EMS_Flags_Byte_EMS098") = 098 * Laenge_Data - Laenge_Data + Allg_Offset 
       SmartTags("SDC\DB_SDC_EMS_FLAGS\_EMS_Flags_Byte_EMS099") = 099 * Laenge_Data - Laenge_Data + Allg_Offset    
       SmartTags("SDC\DB_SDC_EMS_FLAGS\_EMS_Flags_Byte_EMS100") = 100 * Laenge_Data - Laenge_Data + Allg_Offset 
       SmartTags("SDC\DB_SDC_EMS_FLAGS\_EMS_Flags_Byte_EMS101") = 101 * Laenge_Data - Laenge_Data + Allg_Offset 
       SmartTags("SDC\DB_SDC_EMS_FLAGS\_EMS_Flags_Byte_EMS102") = 102 * Laenge_Data - Laenge_Data + Allg_Offset 
       SmartTags("SDC\DB_SDC_EMS_FLAGS\_EMS_Flags_Byte_EMS103") = 103 * Laenge_Data - Laenge_Data + Allg_Offset 
       SmartTags("SDC\DB_SDC_EMS_FLAGS\_EMS_Flags_Byte_EMS104") = 104 * Laenge_Data - Laenge_Data + Allg_Offset 
       SmartTags("SDC\DB_SDC_EMS_FLAGS\_EMS_Flags_Byte_EMS105") = 105 * Laenge_Data - Laenge_Data + Allg_Offset 
       SmartTags("SDC\DB_SDC_EMS_FLAGS\_EMS_Flags_Byte_EMS106") = 106 * Laenge_Data - Laenge_Data + Allg_Offset 
       SmartTags("SDC\DB_SDC_EMS_FLAGS\_EMS_Flags_Byte_EMS107") = 107 * Laenge_Data - Laenge_Data + Allg_Offset 
       SmartTags("SDC\DB_SDC_EMS_FLAGS\_EMS_Flags_Byte_EMS108") = 108 * Laenge_Data - Laenge_Data + Allg_Offset 
       SmartTags("SDC\DB_SDC_EMS_FLAGS\_EMS_Flags_Byte_EMS109") = 109 * Laenge_Data - Laenge_Data + Allg_Offset    
       SmartTags("SDC\DB_SDC_EMS_FLAGS\_EMS_Flags_Byte_EMS110") = 110 * Laenge_Data - Laenge_Data + Allg_Offset   
       SmartTags("SDC\DB_SDC_EMS_FLAGS\_EMS_Flags_Byte_EMS111") = 111 * Laenge_Data - Laenge_Data + Allg_Offset     	
       SmartTags("SDC\DB_SDC_EMS_FLAGS\_EMS_Flags_Byte_EMS112") = 112 * Laenge_Data - Laenge_Data + Allg_Offset 
       SmartTags("SDC\DB_SDC_EMS_FLAGS\_EMS_Flags_Byte_EMS113") = 113 * Laenge_Data - Laenge_Data + Allg_Offset 
       SmartTags("SDC\DB_SDC_EMS_FLAGS\_EMS_Flags_Byte_EMS114") = 114 * Laenge_Data - Laenge_Data + Allg_Offset 
       SmartTags("SDC\DB_SDC_EMS_FLAGS\_EMS_Flags_Byte_EMS115") = 115 * Laenge_Data - Laenge_Data + Allg_Offset 
       SmartTags("SDC\DB_SDC_EMS_FLAGS\_EMS_Flags_Byte_EMS116") = 116 * Laenge_Data - Laenge_Data + Allg_Offset     
       SmartTags("SDC\DB_SDC_EMS_FLAGS\_EMS_Flags_Byte_EMS117") = 117 * Laenge_Data - Laenge_Data + Allg_Offset     
       SmartTags("SDC\DB_SDC_EMS_FLAGS\_EMS_Flags_Byte_EMS118") = 118 * Laenge_Data - Laenge_Data + Allg_Offset     
       SmartTags("SDC\DB_SDC_EMS_FLAGS\_EMS_Flags_Byte_EMS119") = 119 * Laenge_Data - Laenge_Data + Allg_Offset     
       SmartTags("SDC\DB_SDC_EMS_FLAGS\_EMS_Flags_Byte_EMS120") = 120 * Laenge_Data - Laenge_Data + Allg_Offset   
       SmartTags("SDC\DB_SDC_EMS_FLAGS\_EMS_Flags_Byte_EMS121") = 121 * Laenge_Data - Laenge_Data + Allg_Offset     	
       SmartTags("SDC\DB_SDC_EMS_FLAGS\_EMS_Flags_Byte_EMS122") = 122 * Laenge_Data - Laenge_Data + Allg_Offset 
       SmartTags("SDC\DB_SDC_EMS_FLAGS\_EMS_Flags_Byte_EMS123") = 123 * Laenge_Data - Laenge_Data + Allg_Offset 
       SmartTags("SDC\DB_SDC_EMS_FLAGS\_EMS_Flags_Byte_EMS124") = 124 * Laenge_Data - Laenge_Data + Allg_Offset 
       SmartTags("SDC\DB_SDC_EMS_FLAGS\_EMS_Flags_Byte_EMS125") = 125 * Laenge_Data - Laenge_Data + Allg_Offset 
       SmartTags("SDC\DB_SDC_EMS_FLAGS\_EMS_Flags_Byte_EMS126") = 126 * Laenge_Data - Laenge_Data + Allg_Offset     
       SmartTags("SDC\DB_SDC_EMS_FLAGS\_EMS_Flags_Byte_EMS127") = 127 * Laenge_Data - Laenge_Data + Allg_Offset     
       SmartTags("SDC\DB_SDC_EMS_FLAGS\_EMS_Flags_Byte_EMS128") = 128 * Laenge_Data - Laenge_Data + Allg_Offset     
       SmartTags("SDC\DB_SDC_EMS_FLAGS\_EMS_Flags_Byte_EMS129") = 129 * Laenge_Data - Laenge_Data + Allg_Offset      
       SmartTags("SDC\DB_SDC_EMS_FLAGS\_EMS_Flags_Byte_EMS130") = 130 * Laenge_Data - Laenge_Data + Allg_Offset   
       SmartTags("SDC\DB_SDC_EMS_FLAGS\_EMS_Flags_Byte_EMS131") = 131 * Laenge_Data - Laenge_Data + Allg_Offset     	
       SmartTags("SDC\DB_SDC_EMS_FLAGS\_EMS_Flags_Byte_EMS132") = 132 * Laenge_Data - Laenge_Data + Allg_Offset 
       SmartTags("SDC\DB_SDC_EMS_FLAGS\_EMS_Flags_Byte_EMS133") = 133 * Laenge_Data - Laenge_Data + Allg_Offset 
       SmartTags("SDC\DB_SDC_EMS_FLAGS\_EMS_Flags_Byte_EMS134") = 134 * Laenge_Data - Laenge_Data + Allg_Offset 
       SmartTags("SDC\DB_SDC_EMS_FLAGS\_EMS_Flags_Byte_EMS135") = 135 * Laenge_Data - Laenge_Data + Allg_Offset 
       SmartTags("SDC\DB_SDC_EMS_FLAGS\_EMS_Flags_Byte_EMS136") = 136 * Laenge_Data - Laenge_Data + Allg_Offset     
       SmartTags("SDC\DB_SDC_EMS_FLAGS\_EMS_Flags_Byte_EMS137") = 137 * Laenge_Data - Laenge_Data + Allg_Offset     
       SmartTags("SDC\DB_SDC_EMS_FLAGS\_EMS_Flags_Byte_EMS138") = 138 * Laenge_Data - Laenge_Data + Allg_Offset     
       SmartTags("SDC\DB_SDC_EMS_FLAGS\_EMS_Flags_Byte_EMS139") = 139 * Laenge_Data - Laenge_Data + Allg_Offset  
       SmartTags("SDC\DB_SDC_EMS_FLAGS\_EMS_Flags_Byte_EMS140") = 140 * Laenge_Data - Laenge_Data + Allg_Offset   
       SmartTags("SDC\DB_SDC_EMS_FLAGS\_EMS_Flags_Byte_EMS141") = 141 * Laenge_Data - Laenge_Data + Allg_Offset     	
       SmartTags("SDC\DB_SDC_EMS_FLAGS\_EMS_Flags_Byte_EMS142") = 142 * Laenge_Data - Laenge_Data + Allg_Offset 
       SmartTags("SDC\DB_SDC_EMS_FLAGS\_EMS_Flags_Byte_EMS143") = 143 * Laenge_Data - Laenge_Data + Allg_Offset 
       SmartTags("SDC\DB_SDC_EMS_FLAGS\_EMS_Flags_Byte_EMS144") = 144 * Laenge_Data - Laenge_Data + Allg_Offset 
       SmartTags("SDC\DB_SDC_EMS_FLAGS\_EMS_Flags_Byte_EMS145") = 145 * Laenge_Data - Laenge_Data + Allg_Offset 
       SmartTags("SDC\DB_SDC_EMS_FLAGS\_EMS_Flags_Byte_EMS146") = 146 * Laenge_Data - Laenge_Data + Allg_Offset     
       SmartTags("SDC\DB_SDC_EMS_FLAGS\_EMS_Flags_Byte_EMS147") = 147 * Laenge_Data - Laenge_Data + Allg_Offset     
       SmartTags("SDC\DB_SDC_EMS_FLAGS\_EMS_Flags_Byte_EMS148") = 148 * Laenge_Data - Laenge_Data + Allg_Offset     
       SmartTags("SDC\DB_SDC_EMS_FLAGS\_EMS_Flags_Byte_EMS149") = 149 * Laenge_Data - Laenge_Data + Allg_Offset      
       SmartTags("SDC\DB_SDC_EMS_FLAGS\_EMS_Flags_Byte_EMS150") = 150 * Laenge_Data - Laenge_Data + Allg_Offset   
       SmartTags("SDC\DB_SDC_EMS_FLAGS\_EMS_Flags_Byte_EMS151") = 151 * Laenge_Data - Laenge_Data + Allg_Offset     	
       SmartTags("SDC\DB_SDC_EMS_FLAGS\_EMS_Flags_Byte_EMS152") = 152 * Laenge_Data - Laenge_Data + Allg_Offset 
       SmartTags("SDC\DB_SDC_EMS_FLAGS\_EMS_Flags_Byte_EMS153") = 153 * Laenge_Data - Laenge_Data + Allg_Offset 
       SmartTags("SDC\DB_SDC_EMS_FLAGS\_EMS_Flags_Byte_EMS154") = 154 * Laenge_Data - Laenge_Data + Allg_Offset 
       SmartTags("SDC\DB_SDC_EMS_FLAGS\_EMS_Flags_Byte_EMS155") = 155 * Laenge_Data - Laenge_Data + Allg_Offset 
       SmartTags("SDC\DB_SDC_EMS_FLAGS\_EMS_Flags_Byte_EMS156") = 156 * Laenge_Data - Laenge_Data + Allg_Offset     
       SmartTags("SDC\DB_SDC_EMS_FLAGS\_EMS_Flags_Byte_EMS157") = 157 * Laenge_Data - Laenge_Data + Allg_Offset     
       SmartTags("SDC\DB_SDC_EMS_FLAGS\_EMS_Flags_Byte_EMS158") = 158 * Laenge_Data - Laenge_Data + Allg_Offset     
       SmartTags("SDC\DB_SDC_EMS_FLAGS\_EMS_Flags_Byte_EMS159") = 159 * Laenge_Data - Laenge_Data + Allg_Offset      
       SmartTags("SDC\DB_SDC_EMS_FLAGS\_EMS_Flags_Byte_EMS160") = 160 * Laenge_Data - Laenge_Data + Allg_Offset   
       SmartTags("SDC\DB_SDC_EMS_FLAGS\_EMS_Flags_Byte_EMS161") = 161 * Laenge_Data - Laenge_Data + Allg_Offset     	
       SmartTags("SDC\DB_SDC_EMS_FLAGS\_EMS_Flags_Byte_EMS162") = 162 * Laenge_Data - Laenge_Data + Allg_Offset 
       SmartTags("SDC\DB_SDC_EMS_FLAGS\_EMS_Flags_Byte_EMS163") = 163 * Laenge_Data - Laenge_Data + Allg_Offset 
       SmartTags("SDC\DB_SDC_EMS_FLAGS\_EMS_Flags_Byte_EMS164") = 164 * Laenge_Data - Laenge_Data + Allg_Offset 
       SmartTags("SDC\DB_SDC_EMS_FLAGS\_EMS_Flags_Byte_EMS165") = 165 * Laenge_Data - Laenge_Data + Allg_Offset 
       SmartTags("SDC\DB_SDC_EMS_FLAGS\_EMS_Flags_Byte_EMS166") = 166 * Laenge_Data - Laenge_Data + Allg_Offset     
       SmartTags("SDC\DB_SDC_EMS_FLAGS\_EMS_Flags_Byte_EMS167") = 167 * Laenge_Data - Laenge_Data + Allg_Offset     
       SmartTags("SDC\DB_SDC_EMS_FLAGS\_EMS_Flags_Byte_EMS168") = 168 * Laenge_Data - Laenge_Data + Allg_Offset     
       SmartTags("SDC\DB_SDC_EMS_FLAGS\_EMS_Flags_Byte_EMS169") = 169 * Laenge_Data - Laenge_Data + Allg_Offset      
       SmartTags("SDC\DB_SDC_EMS_FLAGS\_EMS_Flags_Byte_EMS170") = 170 * Laenge_Data - Laenge_Data + Allg_Offset   
       SmartTags("SDC\DB_SDC_EMS_FLAGS\_EMS_Flags_Byte_EMS171") = 171 * Laenge_Data - Laenge_Data + Allg_Offset     	
       SmartTags("SDC\DB_SDC_EMS_FLAGS\_EMS_Flags_Byte_EMS172") = 172 * Laenge_Data - Laenge_Data + Allg_Offset 
       SmartTags("SDC\DB_SDC_EMS_FLAGS\_EMS_Flags_Byte_EMS173") = 173 * Laenge_Data - Laenge_Data + Allg_Offset 
       SmartTags("SDC\DB_SDC_EMS_FLAGS\_EMS_Flags_Byte_EMS174") = 174 * Laenge_Data - Laenge_Data + Allg_Offset 
       SmartTags("SDC\DB_SDC_EMS_FLAGS\_EMS_Flags_Byte_EMS175") = 175 * Laenge_Data - Laenge_Data + Allg_Offset 
       SmartTags("SDC\DB_SDC_EMS_FLAGS\_EMS_Flags_Byte_EMS176") = 176 * Laenge_Data - Laenge_Data + Allg_Offset     
       SmartTags("SDC\DB_SDC_EMS_FLAGS\_EMS_Flags_Byte_EMS177") = 177 * Laenge_Data - Laenge_Data + Allg_Offset     
       SmartTags("SDC\DB_SDC_EMS_FLAGS\_EMS_Flags_Byte_EMS178") = 178 * Laenge_Data - Laenge_Data + Allg_Offset     
       SmartTags("SDC\DB_SDC_EMS_FLAGS\_EMS_Flags_Byte_EMS179") = 179 * Laenge_Data - Laenge_Data + Allg_Offset      
       SmartTags("SDC\DB_SDC_EMS_FLAGS\_EMS_Flags_Byte_EMS180") = 180 * Laenge_Data - Laenge_Data + Allg_Offset   
       SmartTags("SDC\DB_SDC_EMS_FLAGS\_EMS_Flags_Byte_EMS181") = 181 * Laenge_Data - Laenge_Data + Allg_Offset     	
       SmartTags("SDC\DB_SDC_EMS_FLAGS\_EMS_Flags_Byte_EMS182") = 182 * Laenge_Data - Laenge_Data + Allg_Offset 
       SmartTags("SDC\DB_SDC_EMS_FLAGS\_EMS_Flags_Byte_EMS183") = 183 * Laenge_Data - Laenge_Data + Allg_Offset 
       SmartTags("SDC\DB_SDC_EMS_FLAGS\_EMS_Flags_Byte_EMS184") = 184 * Laenge_Data - Laenge_Data + Allg_Offset     
       
       
       EMS_Nr = SmartTags("SDC\DB_SDC_EMS_FLAGS\_EMS_Nr")    
       	
